REGION Network 3 (STL)
         L     12288;
         L     "DBIluminaciónMTA".AuxiliarCalculo;
         OW;
         T     "DBIluminaciónMTA".TiempoPANEL;
         NOP   0;
END_REGION

REGION Network 4
   RUNG wire#powerrail
      Contact( "DBIluminaciónMTA".Encendido )
      I_Contact( "DBIluminaciónMTA".AuxiliarEncendidoPermane )
      S_ODT(T_NO := "TLUZ", TV := "DBIluminaciónMTA".TiempoPANEL, R := wire#w1, BI =>, RET_VAL =>)
   END_RUNG
   RUNG wire#powerrail
      I_Contact( "DBIluminaciónMTA".Encendido )
   END_RUNG wire#w1
   // the same network as SCL:
   #_s5time1 := S_ODT(T_NO := "TLUZ",
                      TV := "DBIluminaciónMTA".TiempoPANEL,
                      S := "DBIluminaciónMTA".Encendido AND NOT "DBIluminaciónMTA".AuxiliarEncendidoPermane,
                      R := NOT "DBIluminaciónMTA".Encendido);
END_REGION

REGION Network 5
   RUNG wire#powerrail
      Contact( "TLUZ" )
      S_Coil( #TEMP0 )
   END_RUNG
   // the same network as SCL:
   IF "TLUZ" THEN #TEMP0 := TRUE; END_IF;
END_REGION

REGION Network 6
   RUNG wire#powerrail
      Contact( "Puls.Iluminati" )
      P_Trig( "DBIluminaciónMTA".FLANCOP )
      wire#w1
      I_Contact( "DBIluminaciónMTA".Encendido )
      Coil( "DBIluminaciónMTA".EcendidoPLS )
   END_RUNG
   RUNG wire#powerrail
      Contact( "DBIluminaciónMTA".EcendidoPLS )
   END_RUNG wire#w1
   // the same network as SCL:
   #_w1 := "Puls.Iluminati" AND NOT "DBIluminaciónMTA".FLANCOP;   // rising edge
   "DBIluminaciónMTA".FLANCOP := "Puls.Iluminati";
   "DBIluminaciónMTA".EcendidoPLS := (#_w1 OR "DBIluminaciónMTA".EcendidoPLS) AND NOT "DBIluminaciónMTA".Encendido;
END_REGION

REGION Network 7
   RUNG wire#powerrail
      Contact( "Puls.Iluminati" )
      P_Trig( "DBIluminaciónMTA".FLANCON )
      wire#w1
      Contact( "DBIluminaciónMTA".Encendido )
      Coil( "DBIluminaciónMTA".ApagadoPLS )
   END_RUNG
   RUNG wire#powerrail
      Contact( "DBIluminaciónMTA".ApagadoPLS )
   END_RUNG wire#w1
   // the same network as SCL:
   #_w1 := "Puls.Iluminati" AND NOT "DBIluminaciónMTA".FLANCON;   // rising edge
   "DBIluminaciónMTA".FLANCON := "Puls.Iluminati";
   "DBIluminaciónMTA".ApagadoPLS := (#_w1 OR "DBIluminaciónMTA".ApagadoPLS) AND "DBIluminaciónMTA".Encendido;
END_REGION

REGION Network 8
   "DBIluminaciónMTA".Encendido := "DBIluminaciónMTA".EncendidoPanel OR "DBIluminaciónMTA".MantenerEncendida OR "DBIluminaciónMTA".EcendidoPLS OR ("DBIluminaciónMTA".Encendido AND NOT "DBIluminaciónMTA".ApagadoPanel AND NOT "DBIluminaciónMTA".ApagadoPLS AND NOT #TEMP0 AND NOT "DBIluminaciónMTA".AuxiliarEncendidoPermane) OR ("DBIluminaciónMTA".Encendido AND NOT "DBIluminaciónMTA".AuxiliarEncendidoPermane AND "DBIluminaciónMTA".MantenerEncendida);
END_REGION

REGION Network 9
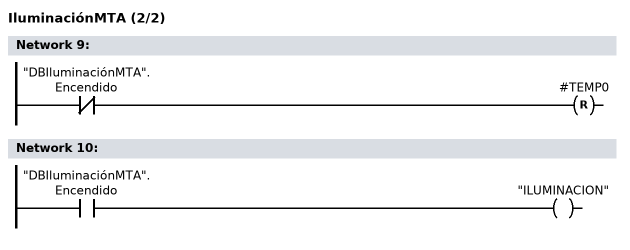
   RUNG wire#powerrail
      I_Contact( "DBIluminaciónMTA".Encendido )
      R_Coil( #TEMP0 )
   END_RUNG
   // the same network as SCL:
   IF NOT "DBIluminaciónMTA".Encendido THEN #TEMP0 := FALSE; END_IF;
END_REGION

REGION Network 10
   RUNG wire#powerrail
      Contact( "DBIluminaciónMTA".Encendido )
      Coil( "ILUMINACION" )
   END_RUNG
   // the same network as SCL:
   "ILUMINACION" := "DBIluminaciónMTA".Encendido;
END_REGION
END_FUNCTION

// folder: OBs de Fallas

ORGANIZATION_BLOCK "OB40"   // OB40, STL
{ S7_Optimized_Access := 'FALSE' }
VERSION : 0.0
BEGIN
END_ORGANIZATION_BLOCK

ORGANIZATION_BLOCK "Cycle Time Fault"   // OB80, STL
{ S7_Optimized_Access := 'FALSE' }
VERSION : 0.0
BEGIN
END_ORGANIZATION_BLOCK

ORGANIZATION_BLOCK "I/O Point Fault 1"   // OB82, LAD
{ S7_Optimized_Access := 'FALSE' }
VERSION : 0.1
BEGIN
END_ORGANIZATION_BLOCK

ORGANIZATION_BLOCK "OB83"   // OB83, STL
{ S7_Optimized_Access := 'FALSE' }
VERSION : 0.1
BEGIN
END_ORGANIZATION_BLOCK

ORGANIZATION_BLOCK "OB Not Loaded Fault"   // OB85, LAD
{ S7_Optimized_Access := 'FALSE' }
VERSION : 0.1
BEGIN
END_ORGANIZATION_BLOCK

ORGANIZATION_BLOCK "Fallo del bastidor"   // OB86, STL
{ S7_Optimized_Access := 'FALSE' }
VERSION : 0.1
BEGIN
END_ORGANIZATION_BLOCK

ORGANIZATION_BLOCK "Communication Fault"   // OB87, LAD
{ S7_Optimized_Access := 'FALSE' }
VERSION : 0.1
BEGIN
END_ORGANIZATION_BLOCK

ORGANIZATION_BLOCK "Complete Restart"   // OB100, LAD
{ S7_Optimized_Access := 'FALSE' }
VERSION : 0.1
BEGIN
END_ORGANIZATION_BLOCK

ORGANIZATION_BLOCK "Programming Error"   // OB121, LAD
{ S7_Optimized_Access := 'FALSE' }
VERSION : 0.1
BEGIN
END_ORGANIZATION_BLOCK

ORGANIZATION_BLOCK "Module Access Error"   // OB122, LAD
{ S7_Optimized_Access := 'FALSE' }
VERSION : 0.1
BEGIN
END_ORGANIZATION_BLOCK

// folder: Panel

FUNCTION_BLOCK "CHControlMotorPanelMTA"   // FB55, LAD
{ S7_Optimized_Access := 'FALSE' }
VERSION : 0.1
   VAR_TEMP   // added for the SCL form of the ladder/FBD networks
      _w1 : Bool;
   END_VAR
BEGIN

REGION Network 1
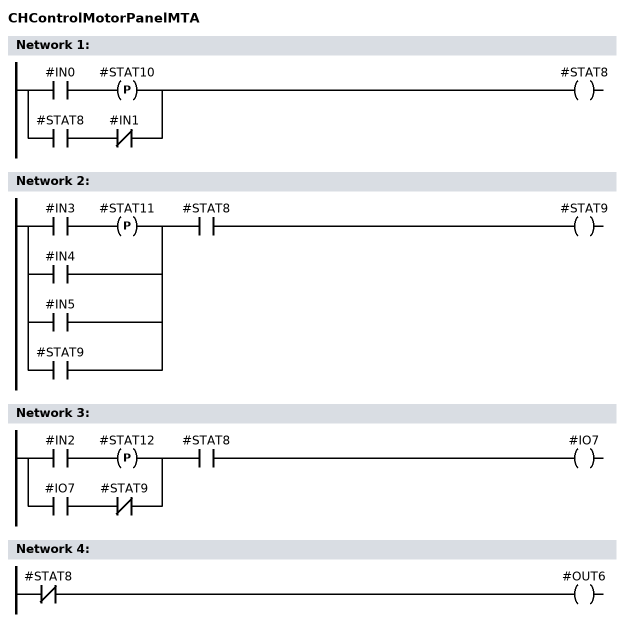
   RUNG wire#powerrail
      Contact( #IN0 )
      P_Trig( #STAT10 )
      wire#w1
      Coil( #STAT8 )
   END_RUNG
   RUNG wire#powerrail
      Contact( #STAT8 )
      I_Contact( #IN1 )
   END_RUNG wire#w1
   // the same network as SCL:
   #_w1 := #IN0 AND NOT #STAT10;   // rising edge
   #STAT10 := #IN0;
   #STAT8 := #_w1 OR (#STAT8 AND NOT #IN1);
END_REGION

REGION Network 2
   RUNG wire#powerrail
      Contact( #IN3 )
      P_Trig( #STAT11 )
      wire#w1
      Contact( #STAT8 )
      Coil( #STAT9 )
   END_RUNG
   RUNG wire#powerrail
      Contact( #IN4 )
   END_RUNG wire#w1
   RUNG wire#powerrail
      Contact( #IN5 )
   END_RUNG wire#w1
   RUNG wire#powerrail
      Contact( #STAT9 )
   END_RUNG wire#w1
   // the same network as SCL:
   #_w1 := #IN3 AND NOT #STAT11;   // rising edge
   #STAT11 := #IN3;
   #STAT9 := (#_w1 OR #IN4 OR #IN5 OR #STAT9) AND #STAT8;
END_REGION

REGION Network 3
   RUNG wire#powerrail
      Contact( #IN2 )
      P_Trig( #STAT12 )
      wire#w1
      Contact( #STAT8 )
      Coil( #IO7 )
   END_RUNG
   RUNG wire#powerrail
      Contact( #IO7 )
      I_Contact( #STAT9 )
   END_RUNG wire#w1
   // the same network as SCL:
   #_w1 := #IN2 AND NOT #STAT12;   // rising edge
   #STAT12 := #IN2;
   #IO7 := (#_w1 OR (#IO7 AND NOT #STAT9)) AND #STAT8;
END_REGION

REGION Network 4
   RUNG wire#powerrail
      I_Contact( #STAT8 )
      Coil( #OUT6 )
   END_RUNG
   // the same network as SCL:
   #OUT6 := NOT #STAT8;
END_REGION
END_FUNCTION_BLOCK

FUNCTION "AnimaciónMTA" : Void   // FC2, LAD
{ S7_Optimized_Access := 'FALSE' }
VERSION : 0.1
   VAR_TEMP   // added for the SCL form of the ladder/FBD networks
      _w1 : Bool;
      _w2 : Bool;
   END_VAR
BEGIN

REGION Network 1: Indicador Chillers
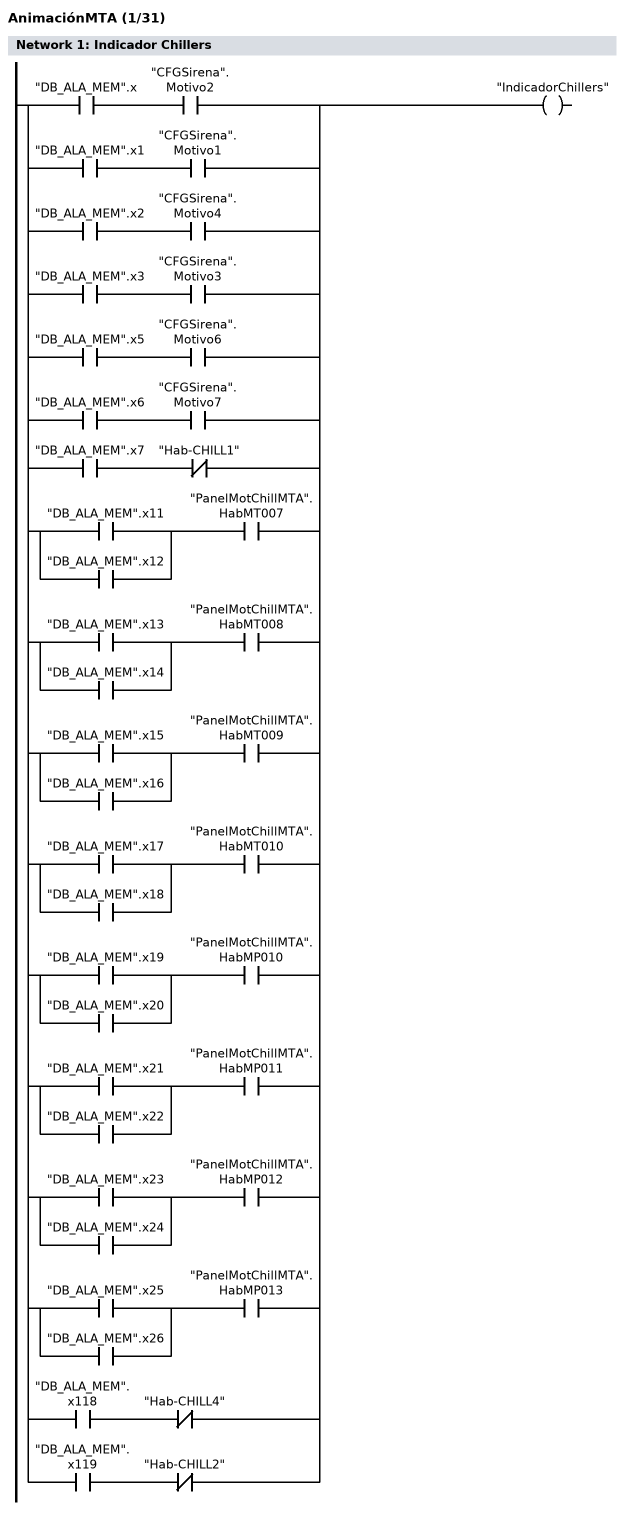
   RUNG wire#powerrail
      Contact( "DB_ALA_MEM".x )
      Contact( "CFGSirena".Motivo2 )
      wire#w1
      Coil( "IndicadorChillers" )
   END_RUNG
   RUNG wire#powerrail
      Contact( "DB_ALA_MEM".x1 )
      Contact( "CFGSirena".Motivo1 )
   END_RUNG wire#w1
   RUNG wire#powerrail
      Contact( "DB_ALA_MEM".x2 )
      Contact( "CFGSirena".Motivo4 )
   END_RUNG wire#w1
   RUNG wire#powerrail
      Contact( "DB_ALA_MEM".x3 )
      Contact( "CFGSirena".Motivo3 )
   END_RUNG wire#w1
   RUNG wire#powerrail
      Contact( "DB_ALA_MEM".x5 )
      Contact( "CFGSirena".Motivo6 )
   END_RUNG wire#w1
   RUNG wire#powerrail
      Contact( "DB_ALA_MEM".x6 )
      Contact( "CFGSirena".Motivo7 )
   END_RUNG wire#w1
   RUNG wire#powerrail
      Contact( "DB_ALA_MEM".x7 )
      I_Contact( "Hab-CHILL1" )
   END_RUNG wire#w1
   RUNG wire#powerrail
      Contact( "DB_ALA_MEM".x11 )
      wire#w2
      Contact( "PanelMotChillMTA".HabMT007 )
   END_RUNG wire#w1
   RUNG wire#powerrail
      Contact( "DB_ALA_MEM".x12 )
   END_RUNG wire#w2
   RUNG wire#powerrail
      Contact( "DB_ALA_MEM".x13 )
      wire#w3
      Contact( "PanelMotChillMTA".HabMT008 )
   END_RUNG wire#w1
   RUNG wire#powerrail
      Contact( "DB_ALA_MEM".x14 )
   END_RUNG wire#w3
   RUNG wire#powerrail
      Contact( "DB_ALA_MEM".x15 )
      wire#w4
      Contact( "PanelMotChillMTA".HabMT009 )
   END_RUNG wire#w1
   RUNG wire#powerrail
      Contact( "DB_ALA_MEM".x16 )
   END_RUNG wire#w4
   RUNG wire#powerrail
      Contact( "DB_ALA_MEM".x17 )
      wire#w5
      Contact( "PanelMotChillMTA".HabMT010 )
   END_RUNG wire#w1
   RUNG wire#powerrail
      Contact( "DB_ALA_MEM".x18 )
   END_RUNG wire#w5
   RUNG wire#powerrail
      Contact( "DB_ALA_MEM".x19 )
      wire#w6
      Contact( "PanelMotChillMTA".HabMP010 )
   END_RUNG wire#w1
   RUNG wire#powerrail
      Contact( "DB_ALA_MEM".x20 )
   END_RUNG wire#w6
   RUNG wire#powerrail
      Contact( "DB_ALA_MEM".x21 )
      wire#w7
      Contact( "PanelMotChillMTA".HabMP011 )
   END_RUNG wire#w1
   RUNG wire#powerrail
      Contact( "DB_ALA_MEM".x22 )
   END_RUNG wire#w7
   RUNG wire#powerrail
      Contact( "DB_ALA_MEM".x23 )
      wire#w8
      Contact( "PanelMotChillMTA".HabMP012 )
   END_RUNG wire#w1
   RUNG wire#powerrail
      Contact( "DB_ALA_MEM".x24 )
   END_RUNG wire#w8
   RUNG wire#powerrail
      Contact( "DB_ALA_MEM".x25 )
      wire#w9
      Contact( "PanelMotChillMTA".HabMP013 )
   END_RUNG wire#w1
   RUNG wire#powerrail
      Contact( "DB_ALA_MEM".x26 )
   END_RUNG wire#w9
   RUNG wire#powerrail
      Contact( "DB_ALA_MEM".x118 )
      I_Contact( "Hab-CHILL4" )
   END_RUNG wire#w1
   RUNG wire#powerrail
      Contact( "DB_ALA_MEM".x119 )
      I_Contact( "Hab-CHILL2" )
   END_RUNG wire#w1
   // the same network as SCL:
   "IndicadorChillers" := ("DB_ALA_MEM".x AND "CFGSirena".Motivo2) OR ("DB_ALA_MEM".x1 AND "CFGSirena".Motivo1) OR ("DB_ALA_MEM".x2 AND "CFGSirena".Motivo4) OR ("DB_ALA_MEM".x3 AND "CFGSirena".Motivo3) OR ("DB_ALA_MEM".x5 AND "CFGSirena".Motivo6) OR ("DB_ALA_MEM".x6 AND "CFGSirena".Motivo7) OR ("DB_ALA_MEM".x7 AND NOT "Hab-CHILL1") OR (("DB_ALA_MEM".x11 OR "DB_ALA_MEM".x12) AND "PanelMotChillMTA".HabMT007) OR (("DB_ALA_MEM".x13 OR "DB_ALA_MEM".x14) AND "PanelMotChillMTA".HabMT008) OR (("DB_ALA_MEM".x15 OR "DB_ALA_MEM".x16) AND "PanelMotChillMTA".HabMT009) OR (("DB_ALA_MEM".x17 OR "DB_ALA_MEM".x18) AND "PanelMotChillMTA".HabMT010) OR (("DB_ALA_MEM".x19 OR "DB_ALA_MEM".x20) AND "PanelMotChillMTA".HabMP010) OR (("DB_ALA_MEM".x21 OR "DB_ALA_MEM".x22) AND "PanelMotChillMTA".HabMP011) OR (("DB_ALA_MEM".x23 OR "DB_ALA_MEM".x24) AND "PanelMotChillMTA".HabMP012) OR (("DB_ALA_MEM".x25 OR "DB_ALA_MEM".x26) AND "PanelMotChillMTA".HabMP013) OR ("DB_ALA_MEM".x118 AND NOT "Hab-CHILL4") OR ("DB_ALA_MEM".x119 AND NOT "Hab-CHILL2");
END_REGION

REGION Network 2: Indicador Torres Chillers
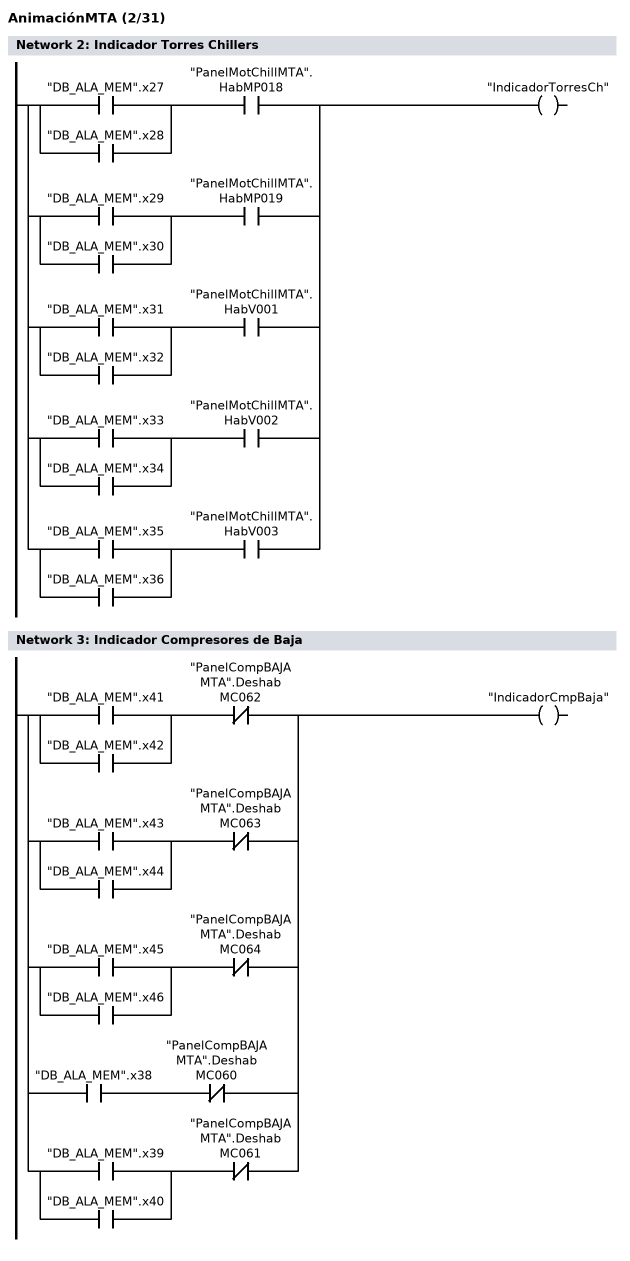
   RUNG wire#powerrail
      Contact( "DB_ALA_MEM".x27 )
      wire#w1
      Contact( "PanelMotChillMTA".HabMP018 )
      wire#w2
      Coil( "IndicadorTorresCh" )
   END_RUNG
   RUNG wire#powerrail
      Contact( "DB_ALA_MEM".x28 )
   END_RUNG wire#w1
   RUNG wire#powerrail
      Contact( "DB_ALA_MEM".x29 )
      wire#w3
      Contact( "PanelMotChillMTA".HabMP019 )
   END_RUNG wire#w2
   RUNG wire#powerrail
      Contact( "DB_ALA_MEM".x30 )
   END_RUNG wire#w3
   RUNG wire#powerrail
      Contact( "DB_ALA_MEM".x31 )
      wire#w4
      Contact( "PanelMotChillMTA".HabV001 )
   END_RUNG wire#w2
   RUNG wire#powerrail
      Contact( "DB_ALA_MEM".x32 )
   END_RUNG wire#w4
   RUNG wire#powerrail
      Contact( "DB_ALA_MEM".x33 )
      wire#w5
      Contact( "PanelMotChillMTA".HabV002 )
   END_RUNG wire#w2
   RUNG wire#powerrail
      Contact( "DB_ALA_MEM".x34 )
   END_RUNG wire#w5
   RUNG wire#powerrail
      Contact( "DB_ALA_MEM".x35 )
      wire#w6
      Contact( "PanelMotChillMTA".HabV003 )
   END_RUNG wire#w2
   RUNG wire#powerrail
      Contact( "DB_ALA_MEM".x36 )
   END_RUNG wire#w6
   // the same network as SCL:
   "IndicadorTorresCh" := (("DB_ALA_MEM".x27 OR "DB_ALA_MEM".x28) AND "PanelMotChillMTA".HabMP018) OR (("DB_ALA_MEM".x29 OR "DB_ALA_MEM".x30) AND "PanelMotChillMTA".HabMP019) OR (("DB_ALA_MEM".x31 OR "DB_ALA_MEM".x32) AND "PanelMotChillMTA".HabV001) OR (("DB_ALA_MEM".x33 OR "DB_ALA_MEM".x34) AND "PanelMotChillMTA".HabV002) OR (("DB_ALA_MEM".x35 OR "DB_ALA_MEM".x36) AND "PanelMotChillMTA".HabV003);
END_REGION

REGION Network 3: Indicador Compresores de Baja
   RUNG wire#powerrail
      Contact( "DB_ALA_MEM".x41 )
      wire#w1
      I_Contact( "PanelCompBAJA MTA".DeshabMC062 )
      wire#w2
      Coil( "IndicadorCmpBaja" )
   END_RUNG
   RUNG wire#powerrail
      Contact( "DB_ALA_MEM".x42 )
   END_RUNG wire#w1
   RUNG wire#powerrail
      Contact( "DB_ALA_MEM".x43 )
      wire#w3
      I_Contact( "PanelCompBAJA MTA".DeshabMC063 )
   END_RUNG wire#w2
   RUNG wire#powerrail
      Contact( "DB_ALA_MEM".x44 )
   END_RUNG wire#w3
   RUNG wire#powerrail
      Contact( "DB_ALA_MEM".x45 )
      wire#w4
      I_Contact( "PanelCompBAJA MTA".DeshabMC064 )
   END_RUNG wire#w2
   RUNG wire#powerrail
      Contact( "DB_ALA_MEM".x46 )
   END_RUNG wire#w4
   RUNG wire#powerrail
      Contact( "DB_ALA_MEM".x38 )
      I_Contact( "PanelCompBAJA MTA".DeshabMC060 )
   END_RUNG wire#w2
   RUNG wire#powerrail
      Contact( "DB_ALA_MEM".x39 )
      wire#w5
      I_Contact( "PanelCompBAJA MTA".DeshabMC061 )
   END_RUNG wire#w2
   RUNG wire#powerrail
      Contact( "DB_ALA_MEM".x40 )
   END_RUNG wire#w5
   // the same network as SCL:
   "IndicadorCmpBaja" := (("DB_ALA_MEM".x41 OR "DB_ALA_MEM".x42) AND NOT "PanelCompBAJA MTA".DeshabMC062) OR (("DB_ALA_MEM".x43 OR "DB_ALA_MEM".x44) AND NOT "PanelCompBAJA MTA".DeshabMC063) OR (("DB_ALA_MEM".x45 OR "DB_ALA_MEM".x46) AND NOT "PanelCompBAJA MTA".DeshabMC064) OR ("DB_ALA_MEM".x38 AND NOT "PanelCompBAJA MTA".DeshabMC060) OR (("DB_ALA_MEM".x39 OR "DB_ALA_MEM".x40) AND NOT "PanelCompBAJA MTA".DeshabMC061);
END_REGION

REGION Network 4: Indicador Secadores de Alta
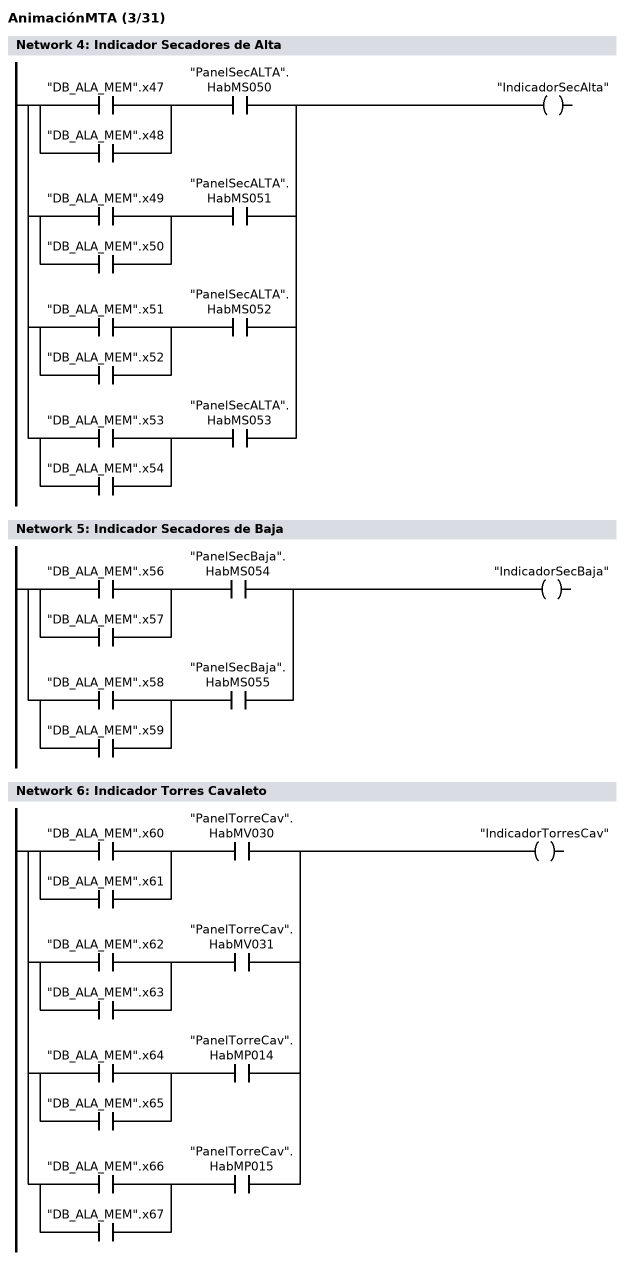
   RUNG wire#powerrail
      Contact( "DB_ALA_MEM".x47 )
      wire#w1
      Contact( "PanelSecALTA".HabMS050 )
      wire#w2
      Coil( "IndicadorSecAlta" )
   END_RUNG
   RUNG wire#powerrail
      Contact( "DB_ALA_MEM".x48 )
   END_RUNG wire#w1
   RUNG wire#powerrail
      Contact( "DB_ALA_MEM".x49 )
      wire#w3
      Contact( "PanelSecALTA".HabMS051 )
   END_RUNG wire#w2
   RUNG wire#powerrail
      Contact( "DB_ALA_MEM".x50 )
   END_RUNG wire#w3
   RUNG wire#powerrail
      Contact( "DB_ALA_MEM".x51 )
      wire#w4
      Contact( "PanelSecALTA".HabMS052 )
   END_RUNG wire#w2
   RUNG wire#powerrail
      Contact( "DB_ALA_MEM".x52 )
   END_RUNG wire#w4
   RUNG wire#powerrail
      Contact( "DB_ALA_MEM".x53 )
      wire#w5
      Contact( "PanelSecALTA".HabMS053 )
   END_RUNG wire#w2
   RUNG wire#powerrail
      Contact( "DB_ALA_MEM".x54 )
   END_RUNG wire#w5
   // the same network as SCL:
   "IndicadorSecAlta" := (("DB_ALA_MEM".x47 OR "DB_ALA_MEM".x48) AND "PanelSecALTA".HabMS050) OR (("DB_ALA_MEM".x49 OR "DB_ALA_MEM".x50) AND "PanelSecALTA".HabMS051) OR (("DB_ALA_MEM".x51 OR "DB_ALA_MEM".x52) AND "PanelSecALTA".HabMS052) OR (("DB_ALA_MEM".x53 OR "DB_ALA_MEM".x54) AND "PanelSecALTA".HabMS053);
END_REGION

REGION Network 5: Indicador Secadores de Baja
   RUNG wire#powerrail
      Contact( "DB_ALA_MEM".x56 )
      wire#w1
      Contact( "PanelSecBaja".HabMS054 )
      wire#w2
      Coil( "IndicadorSecBaja" )
   END_RUNG
   RUNG wire#powerrail
      Contact( "DB_ALA_MEM".x57 )
   END_RUNG wire#w1
   RUNG wire#powerrail
      Contact( "DB_ALA_MEM".x58 )
      wire#w3
      Contact( "PanelSecBaja".HabMS055 )
   END_RUNG wire#w2
   RUNG wire#powerrail
      Contact( "DB_ALA_MEM".x59 )
   END_RUNG wire#w3
   // the same network as SCL:
   "IndicadorSecBaja" := (("DB_ALA_MEM".x56 OR "DB_ALA_MEM".x57) AND "PanelSecBaja".HabMS054) OR (("DB_ALA_MEM".x58 OR "DB_ALA_MEM".x59) AND "PanelSecBaja".HabMS055);
END_REGION

REGION Network 6: Indicador Torres Cavaleto
   RUNG wire#powerrail
      Contact( "DB_ALA_MEM".x60 )
      wire#w1
      Contact( "PanelTorreCav".HabMV030 )
      wire#w2
      Coil( "IndicadorTorresCav" )
   END_RUNG
   RUNG wire#powerrail
      Contact( "DB_ALA_MEM".x61 )
   END_RUNG wire#w1
   RUNG wire#powerrail
      Contact( "DB_ALA_MEM".x62 )
      wire#w3
      Contact( "PanelTorreCav".HabMV031 )
   END_RUNG wire#w2
   RUNG wire#powerrail
      Contact( "DB_ALA_MEM".x63 )
   END_RUNG wire#w3
   RUNG wire#powerrail
      Contact( "DB_ALA_MEM".x64 )
      wire#w4
      Contact( "PanelTorreCav".HabMP014 )
   END_RUNG wire#w2
   RUNG wire#powerrail
      Contact( "DB_ALA_MEM".x65 )
   END_RUNG wire#w4
   RUNG wire#powerrail
      Contact( "DB_ALA_MEM".x66 )
      wire#w5
      Contact( "PanelTorreCav".HabMP015 )
   END_RUNG wire#w2
   RUNG wire#powerrail
      Contact( "DB_ALA_MEM".x67 )
   END_RUNG wire#w5
   // the same network as SCL:
   "IndicadorTorresCav" := (("DB_ALA_MEM".x60 OR "DB_ALA_MEM".x61) AND "PanelTorreCav".HabMV030) OR (("DB_ALA_MEM".x62 OR "DB_ALA_MEM".x63) AND "PanelTorreCav".HabMV031) OR (("DB_ALA_MEM".x64 OR "DB_ALA_MEM".x65) AND "PanelTorreCav".HabMP014) OR (("DB_ALA_MEM".x66 OR "DB_ALA_MEM".x67) AND "PanelTorreCav".HabMP015);
END_REGION

REGION Network 7: Indicador Compresores de Alta
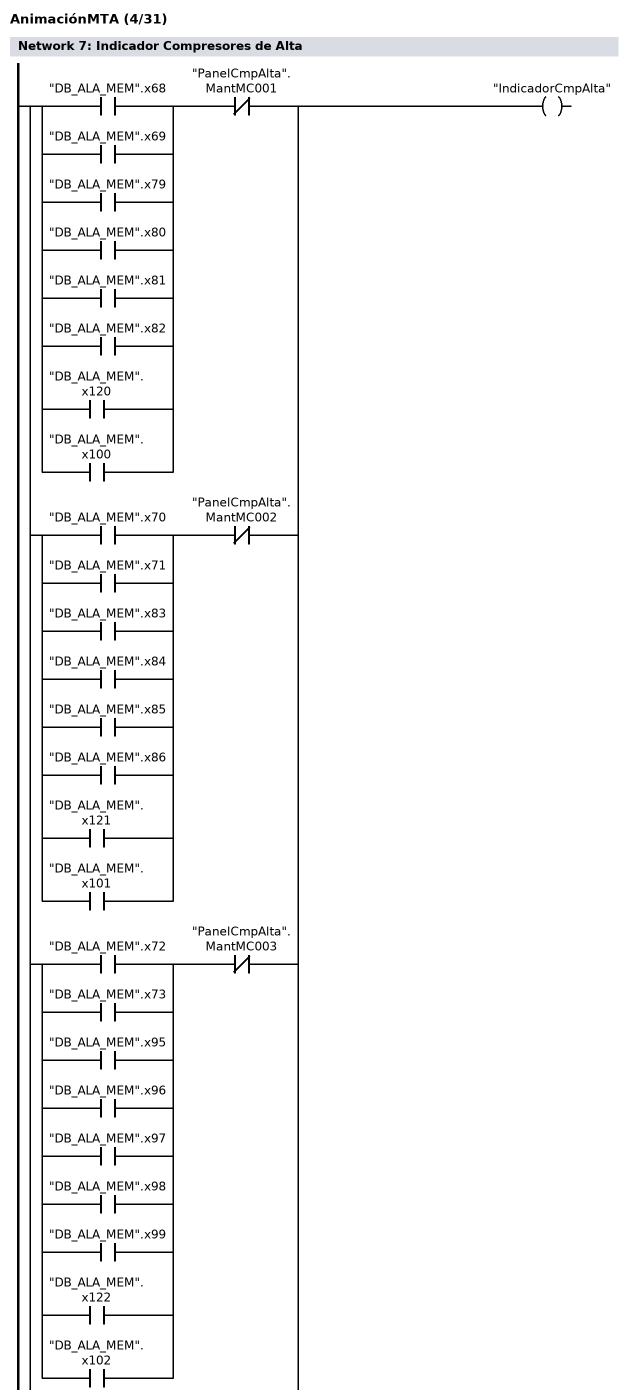
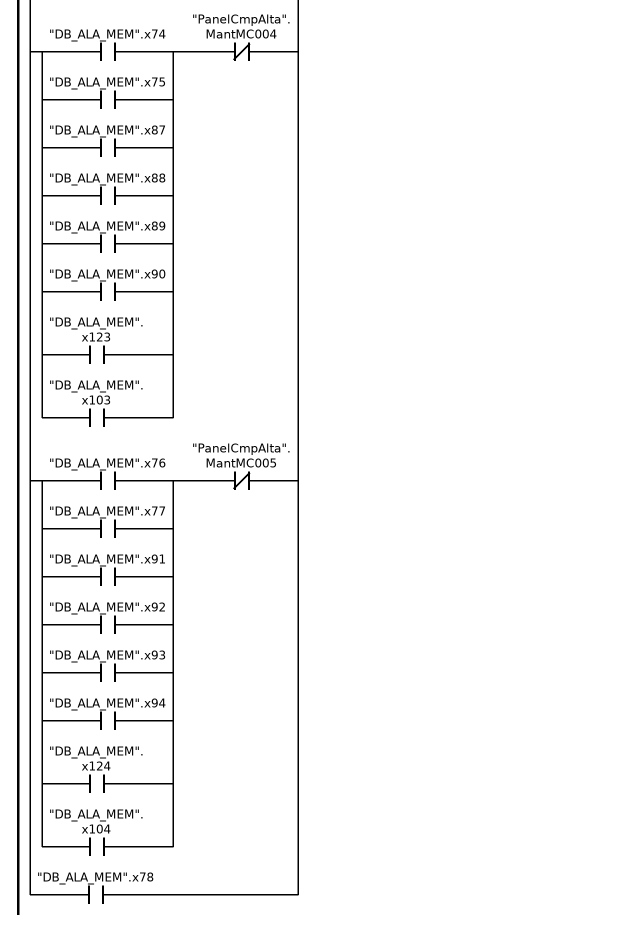
   RUNG wire#powerrail
      Contact( "DB_ALA_MEM".x68 )
      wire#w1
      I_Contact( "PanelCmpAlta".MantMC001 )
      wire#w2
      Coil( "IndicadorCmpAlta" )
   END_RUNG
   RUNG wire#powerrail
      Contact( "DB_ALA_MEM".x69 )
   END_RUNG wire#w1
   RUNG wire#powerrail
      Contact( "DB_ALA_MEM".x79 )
   END_RUNG wire#w1
   RUNG wire#powerrail
      Contact( "DB_ALA_MEM".x80 )
   END_RUNG wire#w1
   RUNG wire#powerrail
      Contact( "DB_ALA_MEM".x81 )
   END_RUNG wire#w1
   RUNG wire#powerrail
      Contact( "DB_ALA_MEM".x82 )
   END_RUNG wire#w1
   RUNG wire#powerrail
      Contact( "DB_ALA_MEM".x120 )
   END_RUNG wire#w1
   RUNG wire#powerrail
      Contact( "DB_ALA_MEM".x100 )
   END_RUNG wire#w1
   RUNG wire#powerrail
      Contact( "DB_ALA_MEM".x70 )
      wire#w3
      I_Contact( "PanelCmpAlta".MantMC002 )
   END_RUNG wire#w2
   RUNG wire#powerrail
      Contact( "DB_ALA_MEM".x71 )
   END_RUNG wire#w3
   RUNG wire#powerrail
      Contact( "DB_ALA_MEM".x83 )
   END_RUNG wire#w3
   RUNG wire#powerrail
      Contact( "DB_ALA_MEM".x84 )
   END_RUNG wire#w3
   RUNG wire#powerrail
      Contact( "DB_ALA_MEM".x85 )
   END_RUNG wire#w3
   RUNG wire#powerrail
      Contact( "DB_ALA_MEM".x86 )
   END_RUNG wire#w3
   RUNG wire#powerrail
      Contact( "DB_ALA_MEM".x121 )
   END_RUNG wire#w3
   RUNG wire#powerrail
      Contact( "DB_ALA_MEM".x101 )
   END_RUNG wire#w3
   RUNG wire#powerrail
      Contact( "DB_ALA_MEM".x72 )
      wire#w4
      I_Contact( "PanelCmpAlta".MantMC003 )
   END_RUNG wire#w2
   RUNG wire#powerrail
      Contact( "DB_ALA_MEM".x73 )
   END_RUNG wire#w4
   RUNG wire#powerrail
      Contact( "DB_ALA_MEM".x95 )
   END_RUNG wire#w4
   RUNG wire#powerrail
      Contact( "DB_ALA_MEM".x96 )
   END_RUNG wire#w4
   RUNG wire#powerrail
      Contact( "DB_ALA_MEM".x97 )
   END_RUNG wire#w4
   RUNG wire#powerrail
      Contact( "DB_ALA_MEM".x98 )
   END_RUNG wire#w4
   RUNG wire#powerrail
      Contact( "DB_ALA_MEM".x99 )
   END_RUNG wire#w4
   RUNG wire#powerrail
      Contact( "DB_ALA_MEM".x122 )
   END_RUNG wire#w4
   RUNG wire#powerrail
      Contact( "DB_ALA_MEM".x102 )
   END_RUNG wire#w4
   RUNG wire#powerrail
      Contact( "DB_ALA_MEM".x74 )
      wire#w5
      I_Contact( "PanelCmpAlta".MantMC004 )
   END_RUNG wire#w2
   RUNG wire#powerrail
      Contact( "DB_ALA_MEM".x75 )
   END_RUNG wire#w5
   RUNG wire#powerrail
      Contact( "DB_ALA_MEM".x87 )
   END_RUNG wire#w5
   RUNG wire#powerrail
      Contact( "DB_ALA_MEM".x88 )
   END_RUNG wire#w5
   RUNG wire#powerrail
      Contact( "DB_ALA_MEM".x89 )
   END_RUNG wire#w5
   RUNG wire#powerrail
      Contact( "DB_ALA_MEM".x90 )
   END_RUNG wire#w5
   RUNG wire#powerrail
      Contact( "DB_ALA_MEM".x123 )
   END_RUNG wire#w5
   RUNG wire#powerrail
      Contact( "DB_ALA_MEM".x103 )
   END_RUNG wire#w5
   RUNG wire#powerrail
      Contact( "DB_ALA_MEM".x76 )
      wire#w6
      I_Contact( "PanelCmpAlta".MantMC005 )
   END_RUNG wire#w2
   RUNG wire#powerrail
      Contact( "DB_ALA_MEM".x77 )
   END_RUNG wire#w6
   RUNG wire#powerrail
      Contact( "DB_ALA_MEM".x91 )
   END_RUNG wire#w6
   RUNG wire#powerrail
      Contact( "DB_ALA_MEM".x92 )
   END_RUNG wire#w6
   RUNG wire#powerrail
      Contact( "DB_ALA_MEM".x93 )
   END_RUNG wire#w6
   RUNG wire#powerrail
      Contact( "DB_ALA_MEM".x94 )
   END_RUNG wire#w6
   RUNG wire#powerrail
      Contact( "DB_ALA_MEM".x124 )
   END_RUNG wire#w6
   RUNG wire#powerrail
      Contact( "DB_ALA_MEM".x104 )
   END_RUNG wire#w6
   RUNG wire#powerrail
      Contact( "DB_ALA_MEM".x78 )
   END_RUNG wire#w2
   // the same network as SCL:
   "IndicadorCmpAlta" := (("DB_ALA_MEM".x68 OR "DB_ALA_MEM".x69 OR "DB_ALA_MEM".x79 OR "DB_ALA_MEM".x80 OR "DB_ALA_MEM".x81 OR "DB_ALA_MEM".x82 OR "DB_ALA_MEM".x120 OR "DB_ALA_MEM".x100) AND NOT "PanelCmpAlta".MantMC001) OR (("DB_ALA_MEM".x70 OR "DB_ALA_MEM".x71 OR "DB_ALA_MEM".x83 OR "DB_ALA_MEM".x84 OR "DB_ALA_MEM".x85 OR "DB_ALA_MEM".x86 OR "DB_ALA_MEM".x121 OR "DB_ALA_MEM".x101) AND NOT "PanelCmpAlta".MantMC002) OR (("DB_ALA_MEM".x72 OR "DB_ALA_MEM".x73 OR "DB_ALA_MEM".x95 OR "DB_ALA_MEM".x96 OR "DB_ALA_MEM".x97 OR "DB_ALA_MEM".x98 OR "DB_ALA_MEM".x99 OR "DB_ALA_MEM".x122 OR "DB_ALA_MEM".x102) AND NOT "PanelCmpAlta".MantMC003) OR (("DB_ALA_MEM".x74 OR "DB_ALA_MEM".x75 OR "DB_ALA_MEM".x87 OR "DB_ALA_MEM".x88 OR "DB_ALA_MEM".x89 OR "DB_ALA_MEM".x90 OR "DB_ALA_MEM".x123 OR "DB_ALA_MEM".x103) AND NOT "PanelCmpAlta".MantMC004) OR (("DB_ALA_MEM".x76 OR "DB_ALA_MEM".x77 OR "DB_ALA_MEM".x91 OR "DB_ALA_MEM".x92 OR "DB_ALA_MEM".x93 OR "DB_ALA_MEM".x94 OR "DB_ALA_MEM".x124 OR "DB_ALA_MEM".x104) AND NOT "PanelCmpAlta".MantMC005) OR "DB_ALA_MEM".x78;
END_REGION

REGION Network 8: Animación MT007 - Bomba Intercambiador LÍNEA 1
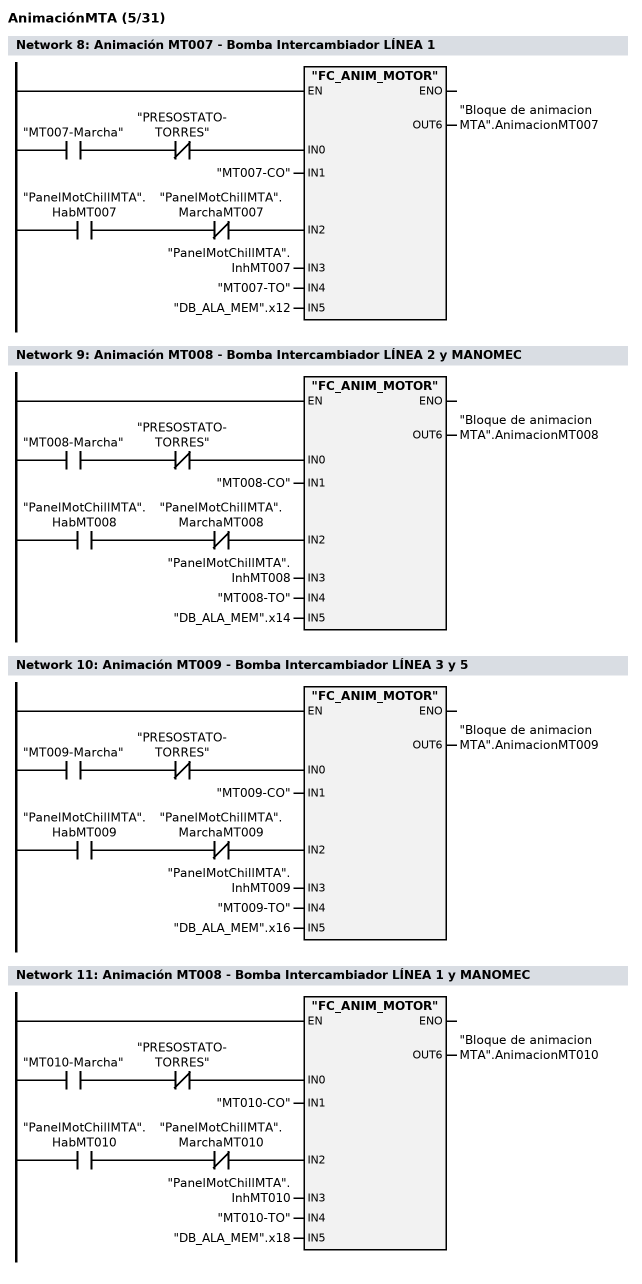
   RUNG wire#powerrail
      "FC_ANIM_MOTOR"(IN0 := wire#w1, IN2 := wire#w2, IN1 := "MT007-CO", IN3 := "PanelMotChillMTA".InhMT007, IN4 := "MT007-TO", IN5 := "DB_ALA_MEM".x12, OUT6 => "Bloque de animacion MTA".AnimacionMT007)
   END_RUNG
   RUNG wire#powerrail
      Contact( "MT007-Marcha" )
      I_Contact( "PRESOSTATO-TORRES" )
   END_RUNG wire#w1
   RUNG wire#powerrail
      Contact( "PanelMotChillMTA".HabMT007 )
      I_Contact( "PanelMotChillMTA".MarchaMT007 )
   END_RUNG wire#w2
   // the same network as SCL:
   "FC_ANIM_MOTOR"(IN0 := "MT007-Marcha" AND NOT "PRESOSTATO-TORRES",
                   IN1 := "MT007-CO",
                   IN2 := "PanelMotChillMTA".HabMT007 AND NOT "PanelMotChillMTA".MarchaMT007,
                   IN3 := "PanelMotChillMTA".InhMT007,
                   IN4 := "MT007-TO",
                   IN5 := "DB_ALA_MEM".x12,
                   OUT6 => "Bloque de animacion MTA".AnimacionMT007);
END_REGION

REGION Network 9: Animación MT008 - Bomba Intercambiador LÍNEA 2 y MANOMEC
   RUNG wire#powerrail
      "FC_ANIM_MOTOR"(IN0 := wire#w1, IN2 := wire#w2, IN1 := "MT008-CO", IN3 := "PanelMotChillMTA".InhMT008, IN4 := "MT008-TO", IN5 := "DB_ALA_MEM".x14, OUT6 => "Bloque de animacion MTA".AnimacionMT008)
   END_RUNG
   RUNG wire#powerrail
      Contact( "MT008-Marcha" )
      I_Contact( "PRESOSTATO-TORRES" )
   END_RUNG wire#w1
   RUNG wire#powerrail
      Contact( "PanelMotChillMTA".HabMT008 )
      I_Contact( "PanelMotChillMTA".MarchaMT008 )
   END_RUNG wire#w2
   // the same network as SCL:
   "FC_ANIM_MOTOR"(IN0 := "MT008-Marcha" AND NOT "PRESOSTATO-TORRES",
                   IN1 := "MT008-CO",
                   IN2 := "PanelMotChillMTA".HabMT008 AND NOT "PanelMotChillMTA".MarchaMT008,
                   IN3 := "PanelMotChillMTA".InhMT008,
                   IN4 := "MT008-TO",
                   IN5 := "DB_ALA_MEM".x14,
                   OUT6 => "Bloque de animacion MTA".AnimacionMT008);
END_REGION

REGION Network 10: Animación MT009 - Bomba Intercambiador LÍNEA 3 y 5
   RUNG wire#powerrail
      "FC_ANIM_MOTOR"(IN0 := wire#w1, IN2 := wire#w2, IN1 := "MT009-CO", IN3 := "PanelMotChillMTA".InhMT009, IN4 := "MT009-TO", IN5 := "DB_ALA_MEM".x16, OUT6 => "Bloque de animacion MTA".AnimacionMT009)
   END_RUNG
   RUNG wire#powerrail
      Contact( "MT009-Marcha" )
      I_Contact( "PRESOSTATO-TORRES" )
   END_RUNG wire#w1
   RUNG wire#powerrail
      Contact( "PanelMotChillMTA".HabMT009 )
      I_Contact( "PanelMotChillMTA".MarchaMT009 )
   END_RUNG wire#w2
   // the same network as SCL:
   "FC_ANIM_MOTOR"(IN0 := "MT009-Marcha" AND NOT "PRESOSTATO-TORRES",
                   IN1 := "MT009-CO",
                   IN2 := "PanelMotChillMTA".HabMT009 AND NOT "PanelMotChillMTA".MarchaMT009,
                   IN3 := "PanelMotChillMTA".InhMT009,
                   IN4 := "MT009-TO",
                   IN5 := "DB_ALA_MEM".x16,
                   OUT6 => "Bloque de animacion MTA".AnimacionMT009);
END_REGION

REGION Network 11: Animación MT008 - Bomba Intercambiador LÍNEA 1 y MANOMEC
   RUNG wire#powerrail
      "FC_ANIM_MOTOR"(IN0 := wire#w1, IN2 := wire#w2, IN1 := "MT010-CO", IN3 := "PanelMotChillMTA".InhMT010, IN4 := "MT010-TO", IN5 := "DB_ALA_MEM".x18, OUT6 => "Bloque de animacion MTA".AnimacionMT010)
   END_RUNG
   RUNG wire#powerrail
      Contact( "MT010-Marcha" )
      I_Contact( "PRESOSTATO-TORRES" )
   END_RUNG wire#w1
   RUNG wire#powerrail
      Contact( "PanelMotChillMTA".HabMT010 )
      I_Contact( "PanelMotChillMTA".MarchaMT010 )
   END_RUNG wire#w2
   // the same network as SCL:
   "FC_ANIM_MOTOR"(IN0 := "MT010-Marcha" AND NOT "PRESOSTATO-TORRES",
                   IN1 := "MT010-CO",
                   IN2 := "PanelMotChillMTA".HabMT010 AND NOT "PanelMotChillMTA".MarchaMT010,
                   IN3 := "PanelMotChillMTA".InhMT010,
                   IN4 := "MT010-TO",
                   IN5 := "DB_ALA_MEM".x18,
                   OUT6 => "Bloque de animacion MTA".AnimacionMT010);
END_REGION

REGION Network 12: Animación MP010 - Bomba Principal Chillers Soplado